// TIA Portal project "ND_PiPl" (V16) (continued)
REGION Network 3: Speicher Stop
   IF (("Schritt_Förderband_Ein" OR "Schritt_Vereinzelner_Ein" OR "Schritt_Horizontalarm_Zurück" OR "Schritt_Vakuum_Ein" OR "Schritt_Vertikalarm_runter" OR "Schritt_Vertikalarm_oben" OR "Schritt_Horizontalarm_vor" OR "Schritt_VertikalarmDeckel_runter" OR "Schritt_Vakuum_aus" OR "Schritt_VertikalarmDeckelweg_oben" OR "Schritt_HorizontalarmDeckel_zurück" OR "Schritt_Vereinzler_aus" OR "Schritt_Zurücksetzten_Anfang") AND "PIPL_Pa_SF_Start") OR ("Deckler_Speicher" AND "PIPL_Pa_SF_Start") OR "Timer_Clean_Reset".Q THEN
       "Stop_Speicher" := FALSE;   // RS flip-flop
   END_IF;
   IF (("Timer_Rückstau".Q AND "PIPL_Pa_SF_ManAuto") OR NOT "PIPL_Pa_SF_Stop" OR "Druck_Zu_Hoch" OR "Druck_Zu_Niedrig") AND ("Schritt_Förderband_Ein" OR "Schritt_Vereinzelner_Ein" OR "Schritt_Horizontalarm_Zurück" OR "Schritt_Vakuum_Ein" OR "Schritt_Vertikalarm_runter" OR "Schritt_Vertikalarm_oben" OR "Schritt_Horizontalarm_vor" OR "Schritt_VertikalarmDeckel_runter" OR "Schritt_Vakuum_aus" OR "Schritt_VertikalarmDeckelweg_oben" OR "Schritt_HorizontalarmDeckel_zurück" OR "Schritt_Vereinzler_aus" OR "Schritt_Zurücksetzten_Anfang") THEN
       "Stop_Speicher" := TRUE;
   END_IF;
END_REGION

REGION Network 4: Wenn keine Deckel vorhanden, dann Vakuum aus
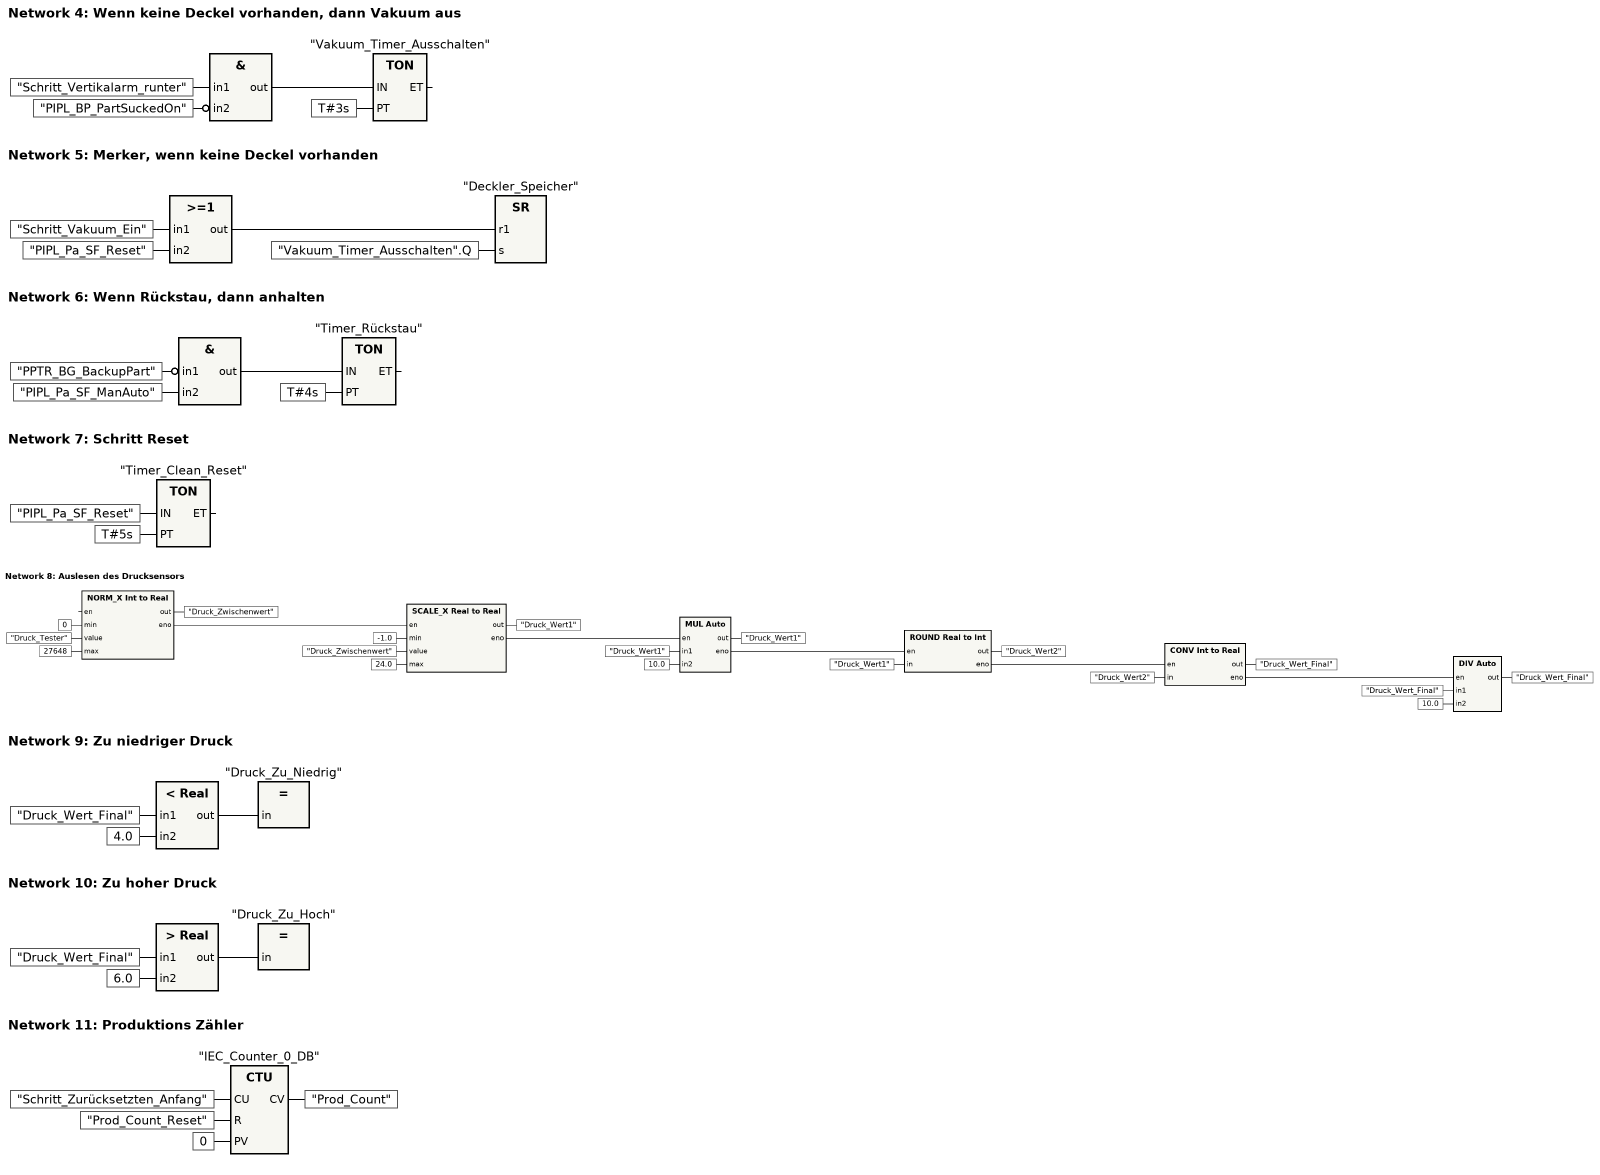
   "Vakuum_Timer_Ausschalten".TON(IN := "Schritt_Vertikalarm_runter" AND NOT "PIPL_BP_PartSuckedOn", PT := T#3s);
END_REGION

REGION Network 5: Merker, wenn keine Deckel vorhanden
   IF "Vakuum_Timer_Ausschalten".Q THEN
       "Deckler_Speicher" := TRUE;   // SR flip-flop
   END_IF;
   IF "Schritt_Vakuum_Ein" OR "PIPL_Pa_SF_Reset" THEN "Deckler_Speicher" := FALSE; END_IF;
END_REGION

REGION Network 6: Wenn Rückstau, dann anhalten
   "Timer_Rückstau".TON(IN := NOT "PPTR_BG_BackupPart" AND "PIPL_Pa_SF_ManAuto", PT := T#4s);
END_REGION

REGION Network 7: Schritt Reset
   "Timer_Clean_Reset".TON(IN := "PIPL_Pa_SF_Reset", PT := T#5s);
END_REGION

REGION Network 8: Auslesen des Drucksensors
   "Druck_Zwischenwert" := NORM_X(MIN := 0, VALUE := "Druck_Tester", MAX := 27648);
   "Druck_Wert1" := SCALE_X(MIN := -1.0, VALUE := "Druck_Zwischenwert", MAX := 24.0);
   "Druck_Wert1" := "Druck_Wert1" * 10.0;
   "Druck_Wert2" := ROUND("Druck_Wert1");
   "Druck_Wert_Final" := INT_TO_REAL("Druck_Wert2");
   "Druck_Wert_Final" := "Druck_Wert_Final" / 10.0;
END_REGION

REGION Network 9: Zu niedriger Druck
   "Druck_Zu_Niedrig" := "Druck_Wert_Final" < 4.0;
END_REGION

REGION Network 10: Zu hoher Druck
   "Druck_Zu_Hoch" := "Druck_Wert_Final" > 6.0;
END_REGION

REGION Network 11: Produktions Zähler
   "IEC_Counter_0_DB".CTU(CU := "Schritt_Zurücksetzten_Anfang",
                          R := "Prod_Count_Reset",
                          PV := 0,
                          CV => "Prod_Count");
END_REGION
END_FUNCTION

FUNCTION "Pick&Place_Manual" : Void   // FC4, FBD
{ S7_Optimized_Access := 'TRUE' }
VERSION : 0.1
BEGIN

REGION Network 1: Eischalten der Maschine
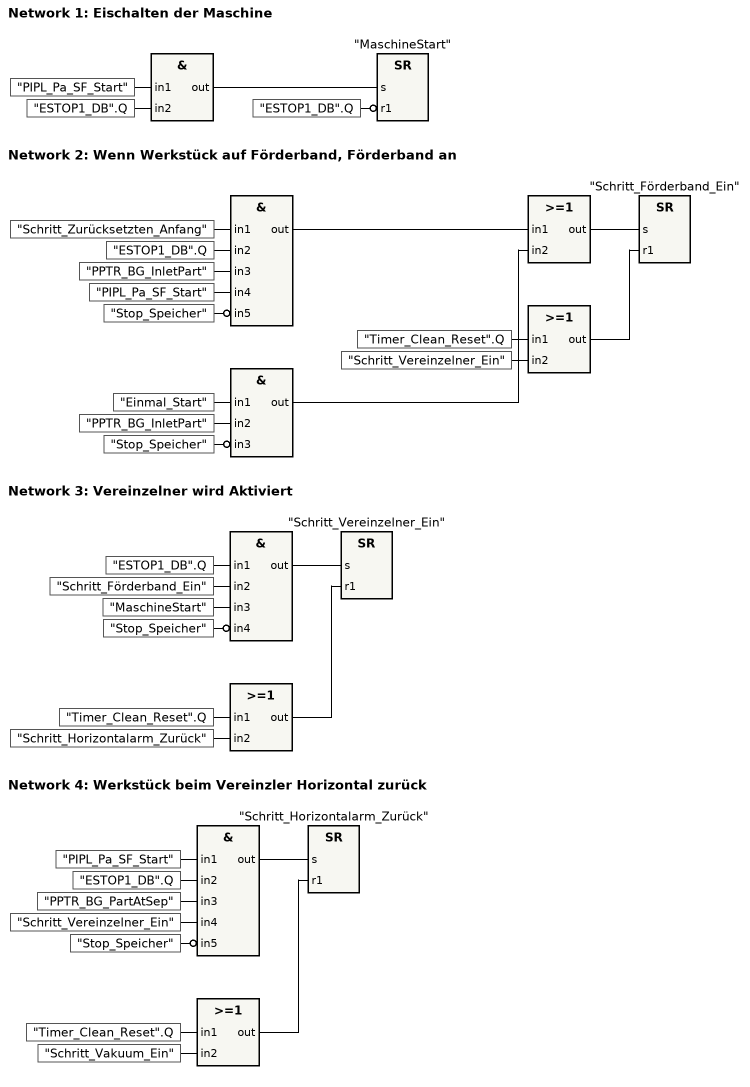
   IF "PIPL_Pa_SF_Start" AND "ESTOP1_DB".Q THEN
       "MaschineStart" := TRUE;   // SR flip-flop
   END_IF;
   IF NOT "ESTOP1_DB".Q THEN "MaschineStart" := FALSE; END_IF;
END_REGION

REGION Network 2: Wenn Werkstück auf Förderband, Förderband an
   IF ("Schritt_Zurücksetzten_Anfang" AND "ESTOP1_DB".Q AND "PPTR_BG_InletPart" AND "PIPL_Pa_SF_Start" AND NOT "Stop_Speicher") OR ("Einmal_Start" AND "PPTR_BG_InletPart" AND NOT "Stop_Speicher") THEN
       "Schritt_Förderband_Ein" := TRUE;   // SR flip-flop
   END_IF;
   IF "Timer_Clean_Reset".Q OR "Schritt_Vereinzelner_Ein" THEN "Schritt_Förderband_Ein" := FALSE; END_IF;
END_REGION

REGION Network 3: Vereinzelner wird Aktiviert
   IF "ESTOP1_DB".Q AND "Schritt_Förderband_Ein" AND "MaschineStart" AND NOT "Stop_Speicher" THEN
       "Schritt_Vereinzelner_Ein" := TRUE;   // SR flip-flop
   END_IF;
   IF "Timer_Clean_Reset".Q OR "Schritt_Horizontalarm_Zurück" THEN
       "Schritt_Vereinzelner_Ein" := FALSE;
   END_IF;
END_REGION

REGION Network 4: Werkstück beim Vereinzler Horizontal zurück
   IF "PIPL_Pa_SF_Start" AND "ESTOP1_DB".Q AND "PPTR_BG_PartAtSep" AND "Schritt_Vereinzelner_Ein" AND NOT "Stop_Speicher" THEN
       "Schritt_Horizontalarm_Zurück" := TRUE;   // SR flip-flop
   END_IF;
   IF "Timer_Clean_Reset".Q OR "Schritt_Vakuum_Ein" THEN "Schritt_Horizontalarm_Zurück" := FALSE; END_IF;
END_REGION

REGION Network 5: Wenn Horizontalarm zurück, Vakuum ein
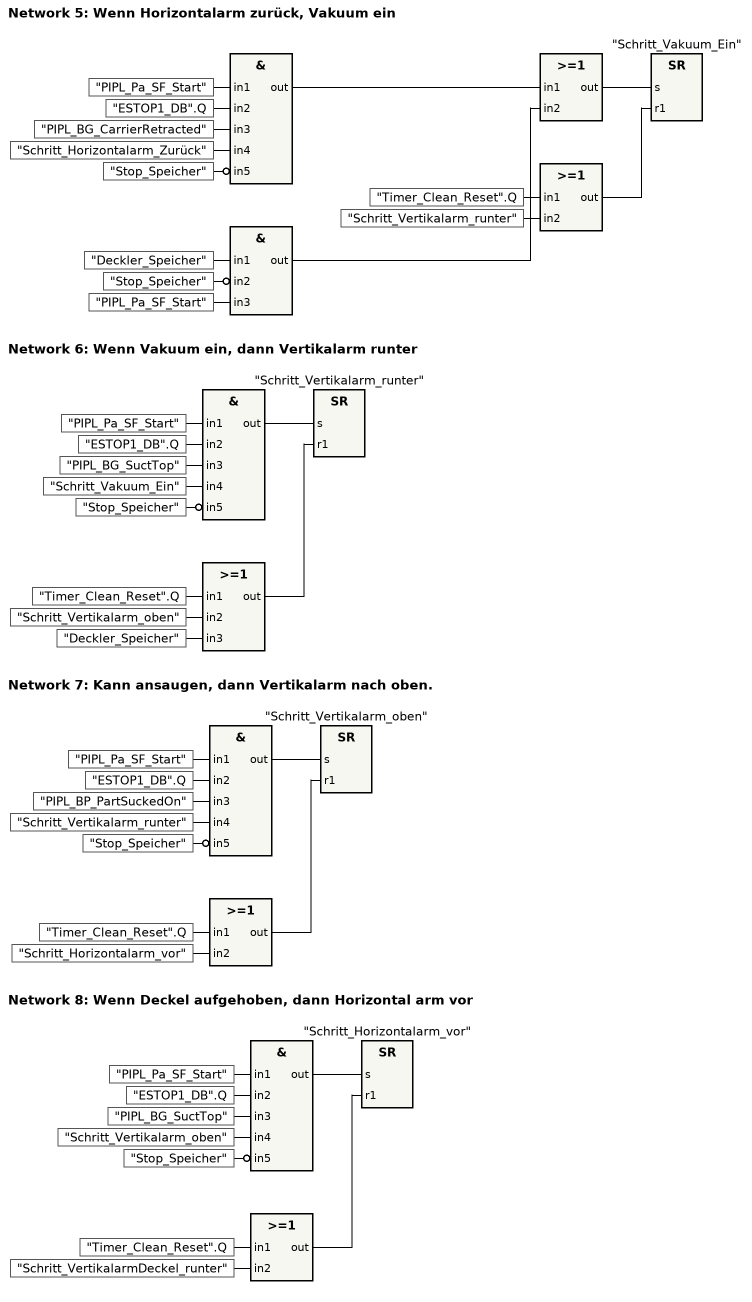
   IF ("PIPL_Pa_SF_Start" AND "ESTOP1_DB".Q AND "PIPL_BG_CarrierRetracted" AND "Schritt_Horizontalarm_Zurück" AND NOT "Stop_Speicher") OR ("Deckler_Speicher" AND NOT "Stop_Speicher" AND "PIPL_Pa_SF_Start") THEN
       "Schritt_Vakuum_Ein" := TRUE;   // SR flip-flop
   END_IF;
   IF "Timer_Clean_Reset".Q OR "Schritt_Vertikalarm_runter" THEN "Schritt_Vakuum_Ein" := FALSE; END_IF;
END_REGION

REGION Network 6: Wenn Vakuum ein, dann Vertikalarm runter
   IF "PIPL_Pa_SF_Start" AND "ESTOP1_DB".Q AND "PIPL_BG_SuctTop" AND "Schritt_Vakuum_Ein" AND NOT "Stop_Speicher" THEN
       "Schritt_Vertikalarm_runter" := TRUE;   // SR flip-flop
   END_IF;
   IF "Timer_Clean_Reset".Q OR "Schritt_Vertikalarm_oben" OR "Deckler_Speicher" THEN
       "Schritt_Vertikalarm_runter" := FALSE;
   END_IF;
END_REGION

REGION Network 7: Kann ansaugen, dann Vertikalarm nach oben.
   IF "PIPL_Pa_SF_Start" AND "ESTOP1_DB".Q AND "PIPL_BP_PartSuckedOn" AND "Schritt_Vertikalarm_runter" AND NOT "Stop_Speicher" THEN
       "Schritt_Vertikalarm_oben" := TRUE;   // SR flip-flop
   END_IF;
   IF "Timer_Clean_Reset".Q OR "Schritt_Horizontalarm_vor" THEN "Schritt_Vertikalarm_oben" := FALSE; END_IF;
END_REGION

REGION Network 8: Wenn Deckel aufgehoben, dann Horizontal arm vor
   IF "PIPL_Pa_SF_Start" AND "ESTOP1_DB".Q AND "PIPL_BG_SuctTop" AND "Schritt_Vertikalarm_oben" AND NOT "Stop_Speicher" THEN
       "Schritt_Horizontalarm_vor" := TRUE;   // SR flip-flop
   END_IF;
   IF "Timer_Clean_Reset".Q OR "Schritt_VertikalarmDeckel_runter" THEN
       "Schritt_Horizontalarm_vor" := FALSE;
   END_IF;
END_REGION

REGION Network 9: Wenn Horizontalarm vor mit Deckel, dann Vertickalarm runter
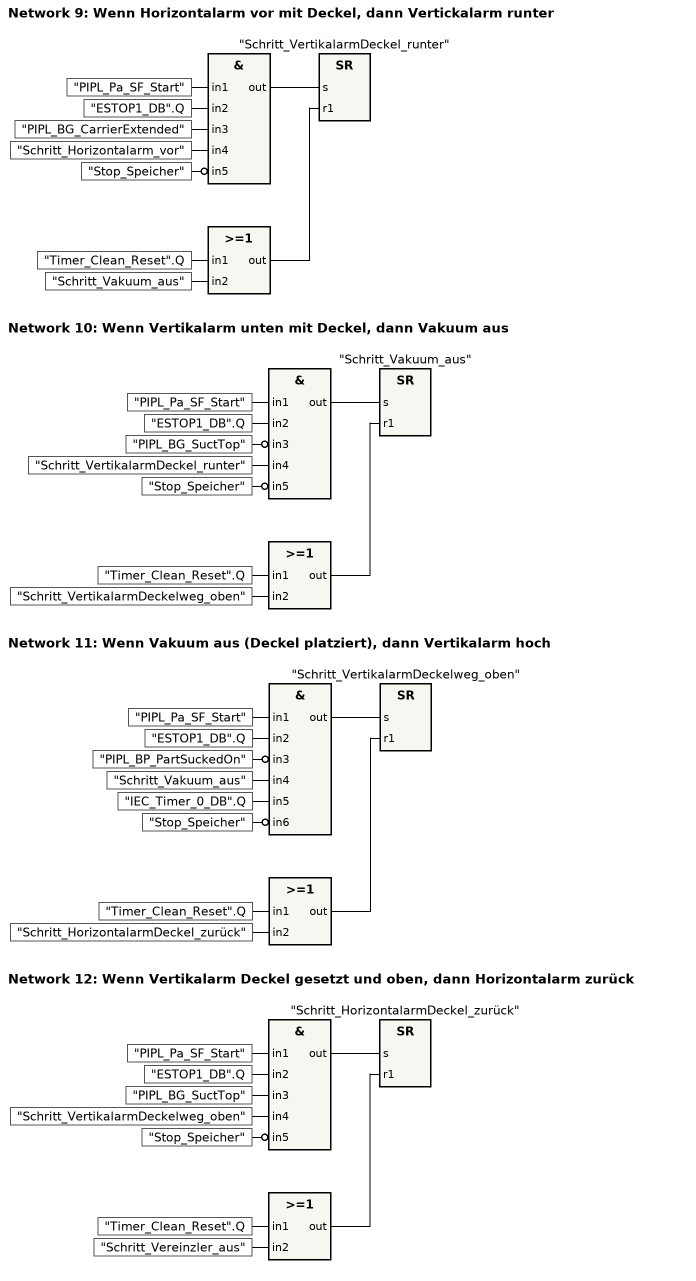
   IF "PIPL_Pa_SF_Start" AND "ESTOP1_DB".Q AND "PIPL_BG_CarrierExtended" AND "Schritt_Horizontalarm_vor" AND NOT "Stop_Speicher" THEN
       "Schritt_VertikalarmDeckel_runter" := TRUE;   // SR flip-flop
   END_IF;
   IF "Timer_Clean_Reset".Q OR "Schritt_Vakuum_aus" THEN "Schritt_VertikalarmDeckel_runter" := FALSE; END_IF;
END_REGION

REGION Network 10: Wenn Vertikalarm unten mit Deckel, dann Vakuum aus
   IF "PIPL_Pa_SF_Start" AND "ESTOP1_DB".Q AND NOT "PIPL_BG_SuctTop" AND "Schritt_VertikalarmDeckel_runter" AND NOT "Stop_Speicher" THEN
       "Schritt_Vakuum_aus" := TRUE;   // SR flip-flop
   END_IF;
   IF "Timer_Clean_Reset".Q OR "Schritt_VertikalarmDeckelweg_oben" THEN
       "Schritt_Vakuum_aus" := FALSE;
   END_IF;
END_REGION

REGION Network 11: Wenn Vakuum aus (Deckel platziert), dann Vertikalarm hoch
   IF "PIPL_Pa_SF_Start" AND "ESTOP1_DB".Q AND NOT "PIPL_BP_PartSuckedOn" AND "Schritt_Vakuum_aus" AND "IEC_Timer_0_DB".Q AND NOT "Stop_Speicher" THEN
       "Schritt_VertikalarmDeckelweg_oben" := TRUE;   // SR flip-flop
   END_IF;
   IF "Timer_Clean_Reset".Q OR "Schritt_HorizontalarmDeckel_zurück" THEN
       "Schritt_VertikalarmDeckelweg_oben" := FALSE;
   END_IF;
END_REGION

REGION Network 12: Wenn Vertikalarm Deckel gesetzt und oben, dann Horizontalarm zurück
   IF "PIPL_Pa_SF_Start" AND "ESTOP1_DB".Q AND "PIPL_BG_SuctTop" AND "Schritt_VertikalarmDeckelweg_oben" AND NOT "Stop_Speicher" THEN
       "Schritt_HorizontalarmDeckel_zurück" := TRUE;   // SR flip-flop
   END_IF;
   IF "Timer_Clean_Reset".Q OR "Schritt_Vereinzler_aus" THEN
       "Schritt_HorizontalarmDeckel_zurück" := FALSE;
   END_IF;
END_REGION

REGION Network 13: Wenn Horizontalarm zurück (Deckel platziert), dann Vereinzler aus
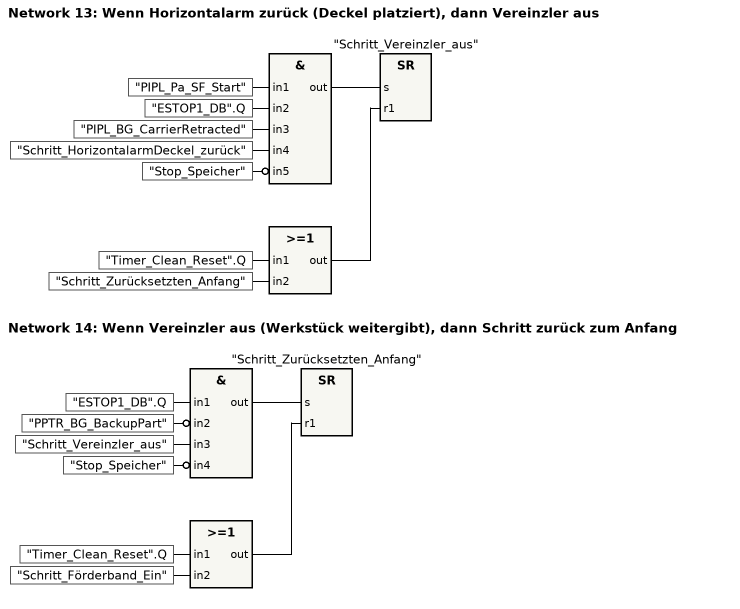
   IF "PIPL_Pa_SF_Start" AND "ESTOP1_DB".Q AND "PIPL_BG_CarrierRetracted" AND "Schritt_HorizontalarmDeckel_zurück" AND NOT "Stop_Speicher" THEN
       "Schritt_Vereinzler_aus" := TRUE;   // SR flip-flop
   END_IF;
   IF "Timer_Clean_Reset".Q OR "Schritt_Zurücksetzten_Anfang" THEN "Schritt_Vereinzler_aus" := FALSE; END_IF;
END_REGION

REGION Network 14: Wenn Vereinzler aus (Werkstück weitergibt), dann Schritt zurück zum Anfang
   IF "ESTOP1_DB".Q AND NOT "PPTR_BG_BackupPart" AND "Schritt_Vereinzler_aus" AND NOT "Stop_Speicher" THEN
       "Schritt_Zurücksetzten_Anfang" := TRUE;   // SR flip-flop
   END_IF;
   IF "Timer_Clean_Reset".Q OR "Schritt_Förderband_Ein" THEN "Schritt_Zurücksetzten_Anfang" := FALSE; END_IF;
END_REGION
END_FUNCTION

FUNCTION "LampenAusgänge_Manual" : Void   // FC5, FBD
{ S7_Optimized_Access := 'TRUE' }
VERSION : 0.1
BEGIN

REGION Network 1: Turmleuchte Grün
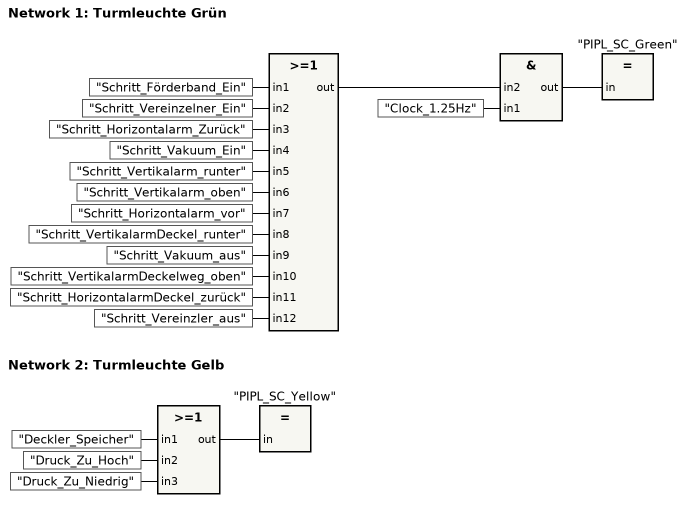
   "PIPL_SC_Green" := ("Schritt_Förderband_Ein" OR "Schritt_Vereinzelner_Ein" OR "Schritt_Horizontalarm_Zurück" OR "Schritt_Vakuum_Ein" OR "Schritt_Vertikalarm_runter" OR "Schritt_Vertikalarm_oben" OR "Schritt_Horizontalarm_vor" OR "Schritt_VertikalarmDeckel_runter" OR "Schritt_Vakuum_aus" OR "Schritt_VertikalarmDeckelweg_oben" OR "Schritt_HorizontalarmDeckel_zurück" OR "Schritt_Vereinzler_aus") AND "Clock_1.25Hz";
END_REGION

REGION Network 2: Turmleuchte Gelb
   "PIPL_SC_Yellow" := "Deckler_Speicher" OR "Druck_Zu_Hoch" OR "Druck_Zu_Niedrig";
END_REGION
END_FUNCTION

FUNCTION "LampenAusgänge_Auto" : Void   // FC6, FBD
{ S7_Optimized_Access := 'TRUE' }
VERSION : 0.1
BEGIN

REGION Network 1: Turmleuchte Grün
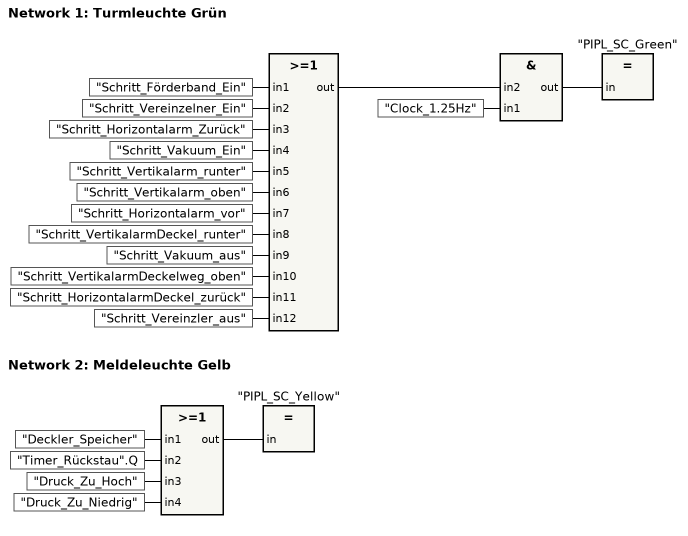
   "PIPL_SC_Green" := ("Schritt_Förderband_Ein" OR "Schritt_Vereinzelner_Ein" OR "Schritt_Horizontalarm_Zurück" OR "Schritt_Vakuum_Ein" OR "Schritt_Vertikalarm_runter" OR "Schritt_Vertikalarm_oben" OR "Schritt_Horizontalarm_vor" OR "Schritt_VertikalarmDeckel_runter" OR "Schritt_Vakuum_aus" OR "Schritt_VertikalarmDeckelweg_oben" OR "Schritt_HorizontalarmDeckel_zurück" OR "Schritt_Vereinzler_aus") AND "Clock_1.25Hz";
END_REGION

REGION Network 2: Meldeleuchte Gelb
   "PIPL_SC_Yellow" := "Deckler_Speicher" OR "Timer_Rückstau".Q OR "Druck_Zu_Hoch" OR "Druck_Zu_Niedrig";
END_REGION
END_FUNCTION

FUNCTION "lampenausgänge_Auto-Manual" : Void   // FC7, FBD
{ S7_Optimized_Access := 'TRUE' }
VERSION : 0.1
BEGIN

REGION Network 1: Turmleuchte Rot
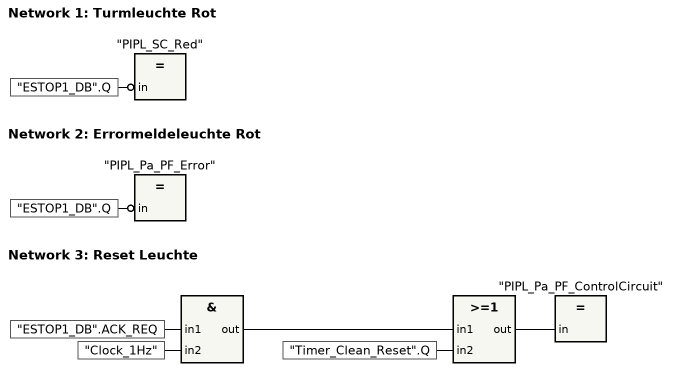
   "PIPL_SC_Red" := NOT "ESTOP1_DB".Q;
END_REGION

REGION Network 2: Errormeldeleuchte Rot
   "PIPL_Pa_PF_Error" := NOT "ESTOP1_DB".Q;
END_REGION

REGION Network 3: Reset Leuchte
   "PIPL_Pa_PF_ControlCircuit" := ("ESTOP1_DB".ACK_REQ AND "Clock_1Hz") OR "Timer_Clean_Reset".Q;
END_REGION

REGION Network 4: Start Taster Lampe
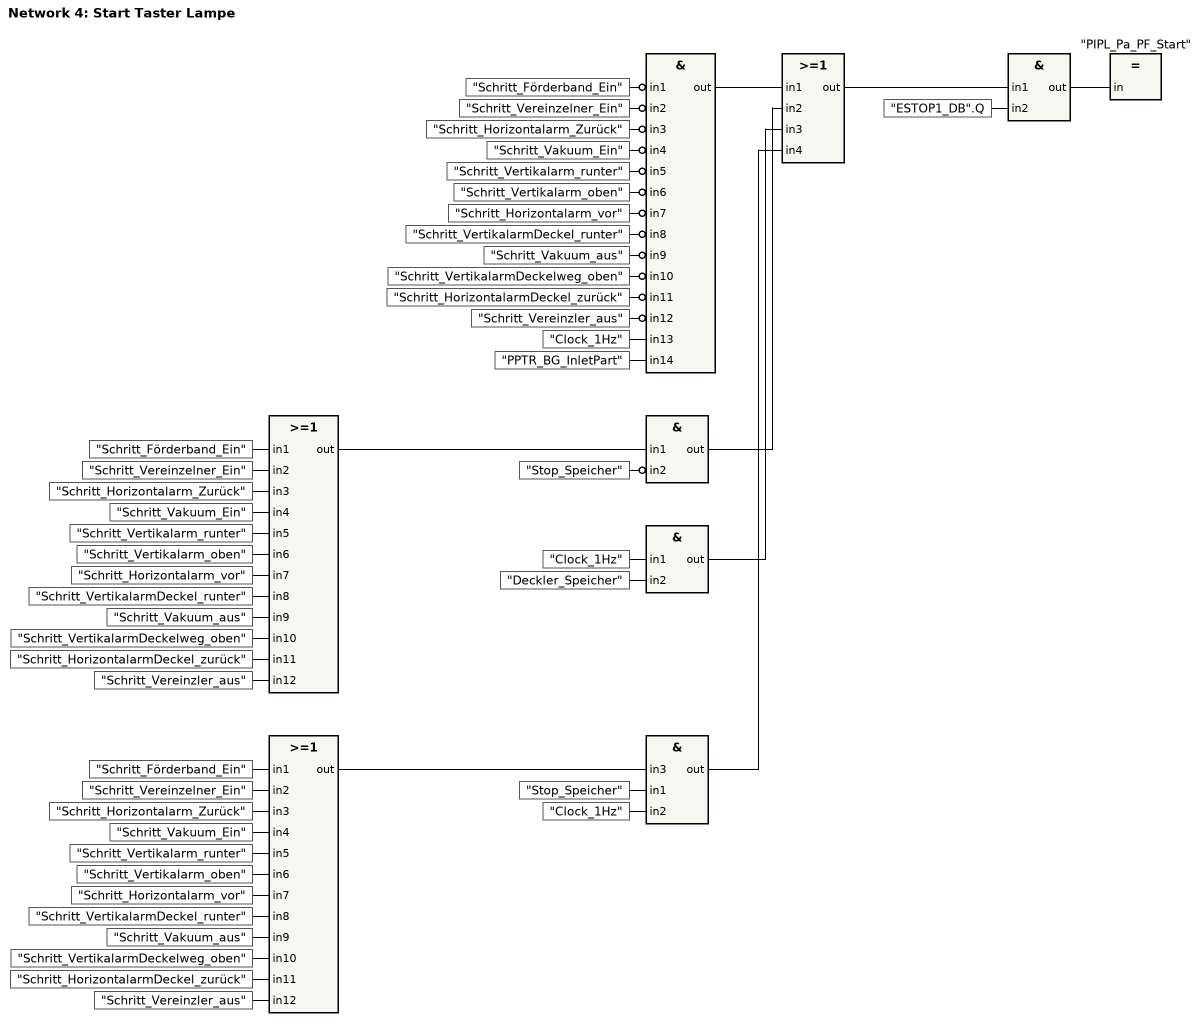
   "PIPL_Pa_PF_Start" := ((NOT "Schritt_Förderband_Ein" AND NOT "Schritt_Vereinzelner_Ein" AND NOT "Schritt_Horizontalarm_Zurück" AND NOT "Schritt_Vakuum_Ein" AND NOT "Schritt_Vertikalarm_runter" AND NOT "Schritt_Vertikalarm_oben" AND NOT "Schritt_Horizontalarm_vor" AND NOT "Schritt_VertikalarmDeckel_runter" AND NOT "Schritt_Vakuum_aus" AND NOT "Schritt_VertikalarmDeckelweg_oben" AND NOT "Schritt_HorizontalarmDeckel_zurück" AND NOT "Schritt_Vereinzler_aus" AND "Clock_1Hz" AND "PPTR_BG_InletPart") OR (("Schritt_Förderband_Ein" OR "Schritt_Vereinzelner_Ein" OR "Schritt_Horizontalarm_Zurück" OR "Schritt_Vakuum_Ein" OR "Schritt_Vertikalarm_runter" OR "Schritt_Vertikalarm_oben" OR "Schritt_Horizontalarm_vor" OR "Schritt_VertikalarmDeckel_runter" OR "Schritt_Vakuum_aus" OR "Schritt_VertikalarmDeckelweg_oben" OR "Schritt_HorizontalarmDeckel_zurück" OR "Schritt_Vereinzler_aus") AND NOT "Stop_Speicher") OR ("Clock_1Hz" AND "Deckler_Speicher") OR (("Schritt_Förderband_Ein" OR "Schritt_Vereinzelner_Ein" OR "Schritt_Horizontalarm_Zurück" OR "Schritt_Vakuum_Ein" OR "Schritt_Vertikalarm_runter" OR "Schritt_Vertikalarm_oben" OR "Schritt_Horizontalarm_vor" OR "Schritt_VertikalarmDeckel_runter" OR "Schritt_Vakuum_aus" OR "Schritt_VertikalarmDeckelweg_oben" OR "Schritt_HorizontalarmDeckel_zurück" OR "Schritt_Vereinzler_aus") AND "Stop_Speicher" AND "Clock_1Hz")) AND "ESTOP1_DB".Q;
END_REGION
END_FUNCTION

FUNCTION "Meldungen_HMI" : Void   // FC8, FBD
{ S7_Optimized_Access := 'TRUE' }
VERSION : 0.1
BEGIN

REGION Network 1: Meldung Not-Aus aktiv
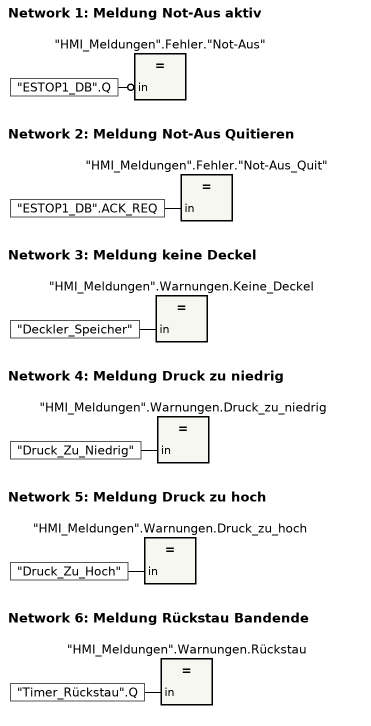
   "HMI_Meldungen".Fehler."Not-Aus" := NOT "ESTOP1_DB".Q;
END_REGION

REGION Network 2: Meldung Not-Aus Quitieren
   "HMI_Meldungen".Fehler."Not-Aus_Quit" := "ESTOP1_DB".ACK_REQ;
END_REGION

REGION Network 3: Meldung keine Deckel
   "HMI_Meldungen".Warnungen.Keine_Deckel := "Deckler_Speicher";
END_REGION

REGION Network 4: Meldung Druck zu niedrig
   "HMI_Meldungen".Warnungen.Druck_zu_niedrig := "Druck_Zu_Niedrig";
END_REGION

REGION Network 5: Meldung Druck zu hoch
   "HMI_Meldungen".Warnungen.Druck_zu_hoch := "Druck_Zu_Hoch";
END_REGION

REGION Network 6: Meldung Rückstau Bandende
   "HMI_Meldungen".Warnungen.Rückstau := "Timer_Rückstau".Q;
END_REGION
END_FUNCTION

ORGANIZATION_BLOCK "Main"   // OB1, FBD, ProgramCycle
TITLE = "Main Program Sweep (Cycle)"
{ S7_Optimized_Access := 'TRUE' }
VERSION : 0.1
   VAR_INPUT
      Initial_Call : Bool;   // Initial call of this OB
      Remanence : Bool;   // =True, if remanent data are available
   END_VAR
BEGIN

REGION Network 1
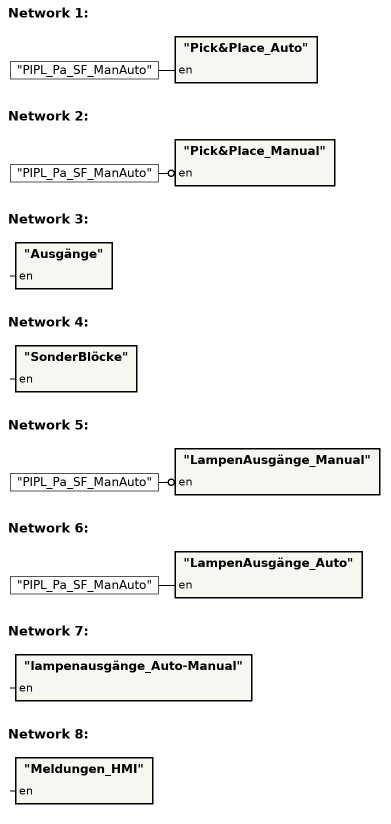
   IF "PIPL_Pa_SF_ManAuto" THEN "Pick&Place_Auto"(); END_IF;
END_REGION

REGION Network 2
   IF NOT "PIPL_Pa_SF_ManAuto" THEN "Pick&Place_Manual"(); END_IF;
END_REGION

REGION Network 3
   "Ausgänge"();
END_REGION

REGION Network 4
   "SonderBlöcke"();
END_REGION

REGION Network 5
   IF NOT "PIPL_Pa_SF_ManAuto" THEN "LampenAusgänge_Manual"(); END_IF;
END_REGION

REGION Network 6
   IF "PIPL_Pa_SF_ManAuto" THEN "LampenAusgänge_Auto"(); END_IF;
END_REGION

REGION Network 7
   "lampenausgänge_Auto-Manual"();
END_REGION

REGION Network 8
   "Meldungen_HMI"();
END_REGION
END_ORGANIZATION_BLOCK

(* ===== HMI "HMI_RT_1" =====
system functions are stored by id; their names below are inferred from use
connection "HMI_1": ETHERNET, S7_1500_OMS

HMI tags "Standard-Variablentabelle"
   "Variable_Bildnummer" : UInt, internal
   "Druck_Wert_Final" : Real = PLC Druck_Wert_Final AT %MD286, 100 ms
   "Prod_Count" : Int = PLC Prod_Count AT %MW1200, 1 s
   "Prod_Count_Reset" : Bool = PLC Prod_Count_Reset AT %M300.0, 1 s

HMI tags "HMI_Meldungen"
   "Fehler" : Word AT %DB120.DBW0, 1 s
   "Meldungen" : Word AT %DB120.DBW2, 1 s
   "Warnungen" : Word AT %DB120.DBW4, 1 s

discrete alarms
   1: 'NOT-AUS Aktiv', class Errors, trigger "Fehler" bit 8
   2: 'NOT-AUS Quitieren', class Errors, trigger "Fehler" bit 9
   3: 'Keine Deckel vorhanden', class Warnings, trigger "Warnungen" bit 10
   4: 'Druck zu niedrig', class Warnings, trigger "Warnungen" bit 8
   5: 'Druck zu hoch', class Warnings, trigger "Warnungen" bit 9
   6: 'Rückstau bandende', class Warnings, trigger "Warnungen" bit 11

text list "Textliste_Bildnamen": 1 'Grundbild'

screen "Start_Bild" 480x272
   GraphicView "Grafikanzeige_1" at 10,7 size 180x55; Picture "PWMA_Logo"
   GraphicView "Grafikanzeige_2" at 295,0 size 185x50; Picture "Pamasol_Zeichen"
   DateTimeField "Datum/Uhrzeit-Feld_1" at 309,57 size 158x21
   Button "Schaltfläche_3" at 0,0 size 473x262; TextOff 'Text'
      on Click: ActivateScreen("DruckAnzeige_Bild", 0)
   Button "Schaltfläche_1" at 30,112 size 188x131; TextOff 'Pamasol Willi Mäder AG Driesbüelstrasse 2 CH-8808 Pfäffikon SZ Schweiz'
   Button "Schaltfläche_4" at 0,0 size 480x270; TextOff '0'
      on Click: ActivateScreen("DruckAnzeige_Bild", 0)
   Button "Schaltfläche_2" at 300,112 size 158x99; TextOff 'Tel. +41 55 417 40 40 Fax. +41 55 417 40 44 info@pamasol.com'
   Softkey "Softkey_F1" at 0,0 size 0x0
      on KeyDown: ActivateScreen("Start_Bild", 0)
   Softkey "Softkey_F2" at 0,0 size 0x0
      on KeyDown: ActivateScreen("DruckAnzeige_Bild", 0)
   Softkey "Softkey_F3" at 0,0 size 0x0
      on KeyDown: ActivateScreen("Ablauf_Meldungen", 0)
   Softkey "Softkey_F4" at 0,0 size 0x0
      on KeyDown: ActivateScreen("Funktions_Bild", 0)

screen "DruckAnzeige_Bild" 480x272
   Softkey "Softkey_F1" at 0,0 size 0x0
      on KeyDown: ActivateScreen("Start_Bild", 0)
   Softkey "Softkey_F2" at 0,0 size 0x0
      on KeyDown: ActivateScreen("DruckAnzeige_Bild", 0)
   DateTimeField "Datum/Uhrzeit-Feld_1" at 312,14 size 158x21
   Gauge "DruckAnzeige" at 243,53 size 176x176; CaptionText 'Pamasol'; UnitText 'Bar'
      ProcessValue <- "Druck_Wert_Final"
   IOField "EA-Feld_1" at 117,99 size 42x28; FormatPattern 9.9
      ProcessValue <- "Druck_Wert_Final"
   TextField "Textfeld_1" at 69,8 size 160x29; Text 'Betriebsdruck'
   Softkey "Softkey_F3" at 0,0 size 0x0
      on KeyDown: ActivateScreen("Ablauf_Meldungen", 0)
   Softkey "Softkey_F4" at 0,0 size 0x0
      on KeyDown: ActivateScreen("Funktions_Bild", 0)

screen "Ablauf_Meldungen" 480x272
   AlarmView "Meldeanzeige_1" at 0,0 size 480x272
   Softkey "Softkey_F1" at 0,0 size 0x0
      on KeyDown: ActivateScreen("Start_Bild", 0)
   Softkey "Softkey_F2" at 0,0 size 0x0
      on KeyDown: ActivateScreen("DruckAnzeige_Bild", 0)
   Softkey "Softkey_F3" at 0,0 size 0x0
      on KeyDown: ActivateScreen("Ablauf_Meldungen", 0)
   Softkey "Softkey_F4" at 0,0 size 0x0
      on KeyDown: ActivateScreen("Funktions_Bild", 0)

screen "Funktions_Bild" 480x272
   Softkey "Softkey_F1" at 0,0 size 0x0
      on KeyDown: ActivateScreen("Start_Bild", 0)
   Softkey "Softkey_F2" at 0,0 size 0x0
      on KeyDown: ActivateScreen("DruckAnzeige_Bild", 0)
   Softkey "Softkey_F3" at 0,0 size 0x0
      on KeyDown: ActivateScreen("Ablauf_Meldungen", 0)
   Softkey "Softkey_F4" at 0,0 size 0x0
      on KeyDown: ActivateScreen("Funktions_Bild", 0)
   IOField "EA-Feld_1" at 215,114 size 51x28; FormatPattern 9999
      ProcessValue <- "Prod_Count"
   Button "Schaltfläche_1" at 184,180 size 112x32; TextOff 'Reset'
      on Press: SetBit("Prod_Count_Reset")
      on Release: ResetBit("Prod_Count_Reset")
   TextField "Textfeld_1" at 127,32 size 226x33; Text 'Produktionsstand'
*)